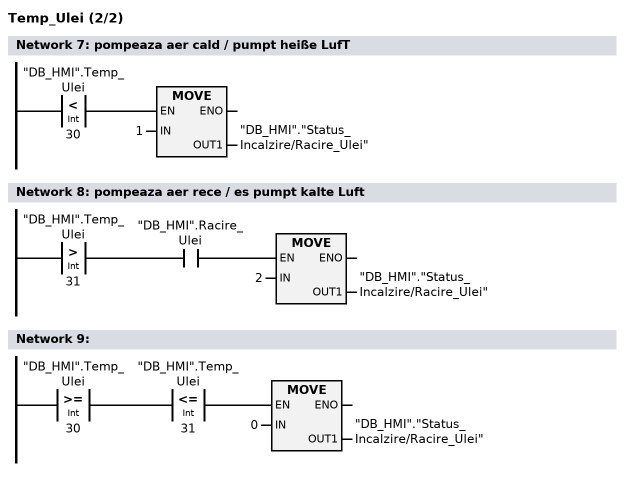
   RUNG wire#powerrail
      { S7_Templates := "SrcType := Int" } LT_Contact(in1 := "DB_HMI".Temp_Ulei, in2 := 30)
      { S7_GenerateENO := "TRUE" } Move(in := 1, out1 => "DB_HMI"."Status_Incalzire/Racire_Ulei")
   END_RUNG
   // the same network as SCL:
   IF "DB_HMI".Temp_Ulei < 30 THEN "DB_HMI"."Status_Incalzire/Racire_Ulei" := 1; END_IF;
END_REGION

REGION Network 8: pompeaza aer rece / es pumpt kalte Luft
   RUNG wire#powerrail
      { S7_Templates := "SrcType := Int" } GT_Contact(in1 := "DB_HMI".Temp_Ulei, in2 := 31)
      Contact( "DB_HMI".Racire_Ulei )
      { S7_GenerateENO := "TRUE" } Move(in := 2, out1 => "DB_HMI"."Status_Incalzire/Racire_Ulei")
   END_RUNG
   // the same network as SCL:
   IF ("DB_HMI".Temp_Ulei > 31) AND "DB_HMI".Racire_Ulei THEN
       "DB_HMI"."Status_Incalzire/Racire_Ulei" := 2;
   END_IF;
END_REGION

REGION Network 9
   RUNG wire#powerrail
      { S7_Templates := "SrcType := Int" } GE_Contact(in1 := "DB_HMI".Temp_Ulei, in2 := 30)
      { S7_Templates := "SrcType := Int" } LE_Contact(in1 := "DB_HMI".Temp_Ulei, in2 := 31)
      { S7_GenerateENO := "TRUE" } Move(in := 0, out1 => "DB_HMI"."Status_Incalzire/Racire_Ulei")
   END_RUNG
   // the same network as SCL:
   IF ("DB_HMI".Temp_Ulei >= 30) AND ("DB_HMI".Temp_Ulei <= 31) THEN
       "DB_HMI"."Status_Incalzire/Racire_Ulei" := 0;
   END_IF;
END_REGION
END_FUNCTION

FUNCTION "Ventilator" : Void   // FC6, LAD
{ S7_Optimized_Access := 'FALSE' }
VERSION : 0.1
BEGIN

REGION Network 1: animatie racire ulei / Ölkühlungsanimation
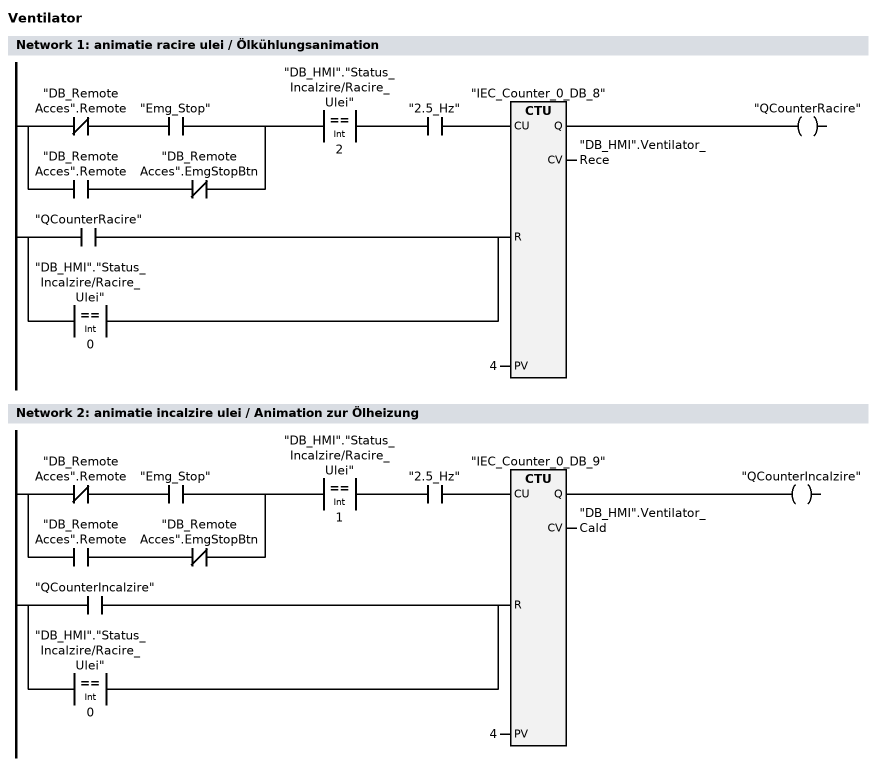
   "IEC_Counter_0_DB_8".CTU(CU := ((NOT "DB_RemoteAcces".Remote AND "Emg_Stop") OR ("DB_RemoteAcces".Remote AND NOT "DB_RemoteAcces".EmgStopBtn)) AND ("DB_HMI"."Status_Incalzire/Racire_Ulei" = 2) AND "2.5_Hz",
                           R := "QCounterRacire" OR ("DB_HMI"."Status_Incalzire/Racire_Ulei" = 0),
                           PV := 4,
                           CV => "DB_HMI".Ventilator_Rece);
   "QCounterRacire" := "IEC_Counter_0_DB_8".Q;
END_REGION

REGION Network 2: animatie incalzire ulei / Animation zur Ölheizung
   "IEC_Counter_0_DB_9".CTU(CU := ((NOT "DB_RemoteAcces".Remote AND "Emg_Stop") OR ("DB_RemoteAcces".Remote AND NOT "DB_RemoteAcces".EmgStopBtn)) AND ("DB_HMI"."Status_Incalzire/Racire_Ulei" = 1) AND "2.5_Hz",
                           R := "QCounterIncalzire" OR ("DB_HMI"."Status_Incalzire/Racire_Ulei" = 0),
                           PV := 4,
                           CV => "DB_HMI".Ventilator_Cald);
   "QCounterIncalzire" := "IEC_Counter_0_DB_9".Q;
END_REGION
END_FUNCTION

FUNCTION "StatusPompe" : Void   // FC19, LAD
{ S7_Optimized_Access := 'FALSE' }
VERSION : 0.1
BEGIN

REGION Network 1
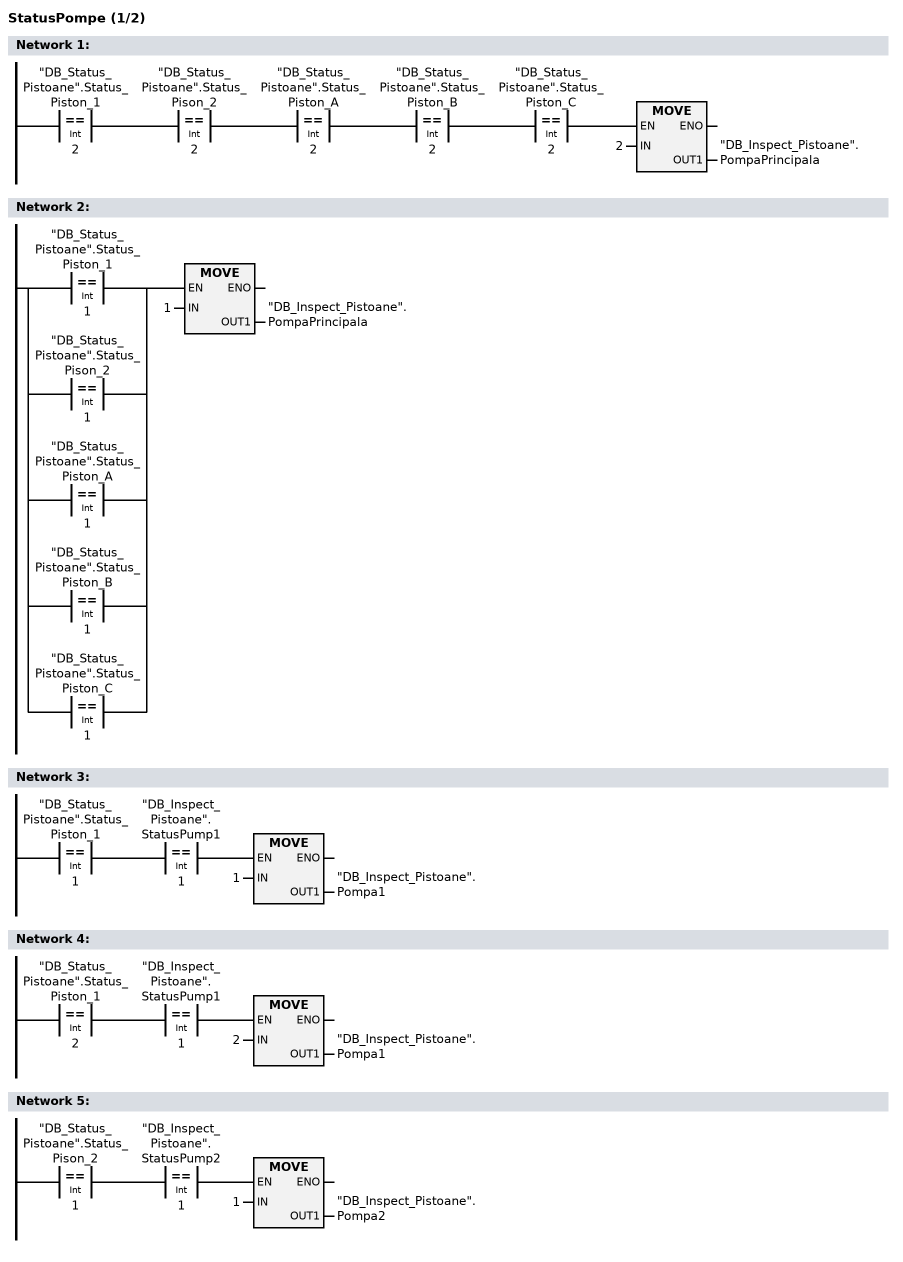
   RUNG wire#powerrail
      { S7_Templates := "SrcType := Int" } EQ_Contact(in1 := "DB_Status_Pistoane".Status_Piston_1, in2 := 2)
      { S7_Templates := "SrcType := Int" } EQ_Contact(in1 := "DB_Status_Pistoane".Status_Pison_2, in2 := 2)
      { S7_Templates := "SrcType := Int" } EQ_Contact(in1 := "DB_Status_Pistoane".Status_Piston_A, in2 := 2)
      { S7_Templates := "SrcType := Int" } EQ_Contact(in1 := "DB_Status_Pistoane".Status_Piston_B, in2 := 2)
      { S7_Templates := "SrcType := Int" } EQ_Contact(in1 := "DB_Status_Pistoane".Status_Piston_C, in2 := 2)
      { S7_GenerateENO := "TRUE" } Move(in := 2, out1 => "DB_Inspect_Pistoane".PompaPrincipala)
   END_RUNG
   // the same network as SCL:
   IF ("DB_Status_Pistoane".Status_Piston_1 = 2) AND ("DB_Status_Pistoane".Status_Pison_2 = 2) AND ("DB_Status_Pistoane".Status_Piston_A = 2) AND ("DB_Status_Pistoane".Status_Piston_B = 2) AND ("DB_Status_Pistoane".Status_Piston_C = 2) THEN
       "DB_Inspect_Pistoane".PompaPrincipala := 2;
   END_IF;
END_REGION

REGION Network 2
   RUNG wire#powerrail
      { S7_Templates := "SrcType := Int" } EQ_Contact(in1 := "DB_Status_Pistoane".Status_Piston_1, in2 := 1)
      wire#w1
      { S7_GenerateENO := "TRUE" } Move(in := 1, out1 => "DB_Inspect_Pistoane".PompaPrincipala)
   END_RUNG
   RUNG wire#powerrail
      { S7_Templates := "SrcType := Int" } EQ_Contact(in1 := "DB_Status_Pistoane".Status_Pison_2, in2 := 1)
   END_RUNG wire#w1
   RUNG wire#powerrail
      { S7_Templates := "SrcType := Int" } EQ_Contact(in1 := "DB_Status_Pistoane".Status_Piston_A, in2 := 1)
   END_RUNG wire#w1
   RUNG wire#powerrail
      { S7_Templates := "SrcType := Int" } EQ_Contact(in1 := "DB_Status_Pistoane".Status_Piston_B, in2 := 1)
   END_RUNG wire#w1
   RUNG wire#powerrail
      { S7_Templates := "SrcType := Int" } EQ_Contact(in1 := "DB_Status_Pistoane".Status_Piston_C, in2 := 1)
   END_RUNG wire#w1
   // the same network as SCL:
   IF ("DB_Status_Pistoane".Status_Piston_1 = 1) OR ("DB_Status_Pistoane".Status_Pison_2 = 1) OR ("DB_Status_Pistoane".Status_Piston_A = 1) OR ("DB_Status_Pistoane".Status_Piston_B = 1) OR ("DB_Status_Pistoane".Status_Piston_C = 1) THEN
       "DB_Inspect_Pistoane".PompaPrincipala := 1;
   END_IF;
END_REGION

REGION Network 3
   RUNG wire#powerrail
      { S7_Templates := "SrcType := Int" } EQ_Contact(in1 := "DB_Status_Pistoane".Status_Piston_1, in2 := 1)
      { S7_Templates := "SrcType := Int" } EQ_Contact(in1 := "DB_Inspect_Pistoane".StatusPump1, in2 := 1)
      { S7_GenerateENO := "TRUE" } Move(in := 1, out1 => "DB_Inspect_Pistoane".Pompa1)
   END_RUNG
   // the same network as SCL:
   IF ("DB_Status_Pistoane".Status_Piston_1 = 1) AND ("DB_Inspect_Pistoane".StatusPump1 = 1) THEN
       "DB_Inspect_Pistoane".Pompa1 := 1;
   END_IF;
END_REGION

REGION Network 4
   RUNG wire#powerrail
      { S7_Templates := "SrcType := Int" } EQ_Contact(in1 := "DB_Status_Pistoane".Status_Piston_1, in2 := 2)
      { S7_Templates := "SrcType := Int" } EQ_Contact(in1 := "DB_Inspect_Pistoane".StatusPump1, in2 := 1)
      { S7_GenerateENO := "TRUE" } Move(in := 2, out1 => "DB_Inspect_Pistoane".Pompa1)
   END_RUNG
   // the same network as SCL:
   IF ("DB_Status_Pistoane".Status_Piston_1 = 2) AND ("DB_Inspect_Pistoane".StatusPump1 = 1) THEN
       "DB_Inspect_Pistoane".Pompa1 := 2;
   END_IF;
END_REGION

REGION Network 5
   RUNG wire#powerrail
      { S7_Templates := "SrcType := Int" } EQ_Contact(in1 := "DB_Status_Pistoane".Status_Pison_2, in2 := 1)
      { S7_Templates := "SrcType := Int" } EQ_Contact(in1 := "DB_Inspect_Pistoane".StatusPump2, in2 := 1)
      { S7_GenerateENO := "TRUE" } Move(in := 1, out1 => "DB_Inspect_Pistoane".Pompa2)
   END_RUNG
   // the same network as SCL:
   IF ("DB_Status_Pistoane".Status_Pison_2 = 1) AND ("DB_Inspect_Pistoane".StatusPump2 = 1) THEN
       "DB_Inspect_Pistoane".Pompa2 := 1;
   END_IF;
END_REGION

REGION Network 6
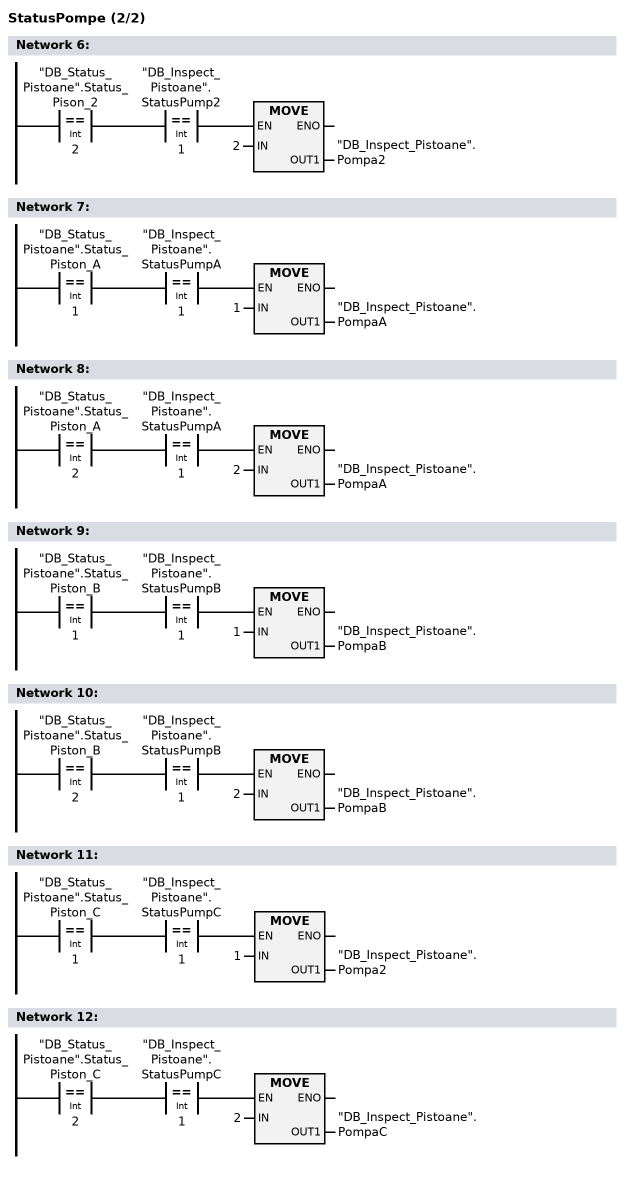
   RUNG wire#powerrail
      { S7_Templates := "SrcType := Int" } EQ_Contact(in1 := "DB_Status_Pistoane".Status_Pison_2, in2 := 2)
      { S7_Templates := "SrcType := Int" } EQ_Contact(in1 := "DB_Inspect_Pistoane".StatusPump2, in2 := 1)
      { S7_GenerateENO := "TRUE" } Move(in := 2, out1 => "DB_Inspect_Pistoane".Pompa2)
   END_RUNG
   // the same network as SCL:
   IF ("DB_Status_Pistoane".Status_Pison_2 = 2) AND ("DB_Inspect_Pistoane".StatusPump2 = 1) THEN
       "DB_Inspect_Pistoane".Pompa2 := 2;
   END_IF;
END_REGION

REGION Network 7
   RUNG wire#powerrail
      { S7_Templates := "SrcType := Int" } EQ_Contact(in1 := "DB_Status_Pistoane".Status_Piston_A, in2 := 1)
      { S7_Templates := "SrcType := Int" } EQ_Contact(in1 := "DB_Inspect_Pistoane".StatusPumpA, in2 := 1)
      { S7_GenerateENO := "TRUE" } Move(in := 1, out1 => "DB_Inspect_Pistoane".PompaA)
   END_RUNG
   // the same network as SCL:
   IF ("DB_Status_Pistoane".Status_Piston_A = 1) AND ("DB_Inspect_Pistoane".StatusPumpA = 1) THEN
       "DB_Inspect_Pistoane".PompaA := 1;
   END_IF;
END_REGION

REGION Network 8
   RUNG wire#powerrail
      { S7_Templates := "SrcType := Int" } EQ_Contact(in1 := "DB_Status_Pistoane".Status_Piston_A, in2 := 2)
      { S7_Templates := "SrcType := Int" } EQ_Contact(in1 := "DB_Inspect_Pistoane".StatusPumpA, in2 := 1)
      { S7_GenerateENO := "TRUE" } Move(in := 2, out1 => "DB_Inspect_Pistoane".PompaA)
   END_RUNG
   // the same network as SCL:
   IF ("DB_Status_Pistoane".Status_Piston_A = 2) AND ("DB_Inspect_Pistoane".StatusPumpA = 1) THEN
       "DB_Inspect_Pistoane".PompaA := 2;
   END_IF;
END_REGION

REGION Network 9
   RUNG wire#powerrail
      { S7_Templates := "SrcType := Int" } EQ_Contact(in1 := "DB_Status_Pistoane".Status_Piston_B, in2 := 1)
      { S7_Templates := "SrcType := Int" } EQ_Contact(in1 := "DB_Inspect_Pistoane".StatusPumpB, in2 := 1)
      { S7_GenerateENO := "TRUE" } Move(in := 1, out1 => "DB_Inspect_Pistoane".PompaB)
   END_RUNG
   // the same network as SCL:
   IF ("DB_Status_Pistoane".Status_Piston_B = 1) AND ("DB_Inspect_Pistoane".StatusPumpB = 1) THEN
       "DB_Inspect_Pistoane".PompaB := 1;
   END_IF;
END_REGION

REGION Network 10
   RUNG wire#powerrail
      { S7_Templates := "SrcType := Int" } EQ_Contact(in1 := "DB_Status_Pistoane".Status_Piston_B, in2 := 2)
      { S7_Templates := "SrcType := Int" } EQ_Contact(in1 := "DB_Inspect_Pistoane".StatusPumpB, in2 := 1)
      { S7_GenerateENO := "TRUE" } Move(in := 2, out1 => "DB_Inspect_Pistoane".PompaB)
   END_RUNG
   // the same network as SCL:
   IF ("DB_Status_Pistoane".Status_Piston_B = 2) AND ("DB_Inspect_Pistoane".StatusPumpB = 1) THEN
       "DB_Inspect_Pistoane".PompaB := 2;
   END_IF;
END_REGION

REGION Network 11
   RUNG wire#powerrail
      { S7_Templates := "SrcType := Int" } EQ_Contact(in1 := "DB_Status_Pistoane".Status_Piston_C, in2 := 1)
      { S7_Templates := "SrcType := Int" } EQ_Contact(in1 := "DB_Inspect_Pistoane".StatusPumpC, in2 := 1)
      { S7_GenerateENO := "TRUE" } Move(in := 1, out1 => "DB_Inspect_Pistoane".Pompa2)
   END_RUNG
   // the same network as SCL:
   IF ("DB_Status_Pistoane".Status_Piston_C = 1) AND ("DB_Inspect_Pistoane".StatusPumpC = 1) THEN
       "DB_Inspect_Pistoane".Pompa2 := 1;
   END_IF;
END_REGION

REGION Network 12
   RUNG wire#powerrail
      { S7_Templates := "SrcType := Int" } EQ_Contact(in1 := "DB_Status_Pistoane".Status_Piston_C, in2 := 2)
      { S7_Templates := "SrcType := Int" } EQ_Contact(in1 := "DB_Inspect_Pistoane".StatusPumpC, in2 := 1)
      { S7_GenerateENO := "TRUE" } Move(in := 2, out1 => "DB_Inspect_Pistoane".PompaC)
   END_RUNG
   // the same network as SCL:
   IF ("DB_Status_Pistoane".Status_Piston_C = 2) AND ("DB_Inspect_Pistoane".StatusPumpC = 1) THEN
       "DB_Inspect_Pistoane".PompaC := 2;
   END_IF;
END_REGION
END_FUNCTION

// folder: Statie Distribuire/Animatii

FUNCTION_BLOCK "Animatie_Banda_1"   // FB2, LAD
{ S7_Optimized_Access := 'FALSE' }
VERSION : 0.1
   VAR_TEMP   // added for the SCL form of the ladder/FBD networks
      _w1 : Bool;
      _w2 : Bool;
   END_VAR
BEGIN

REGION Network 1: ceva
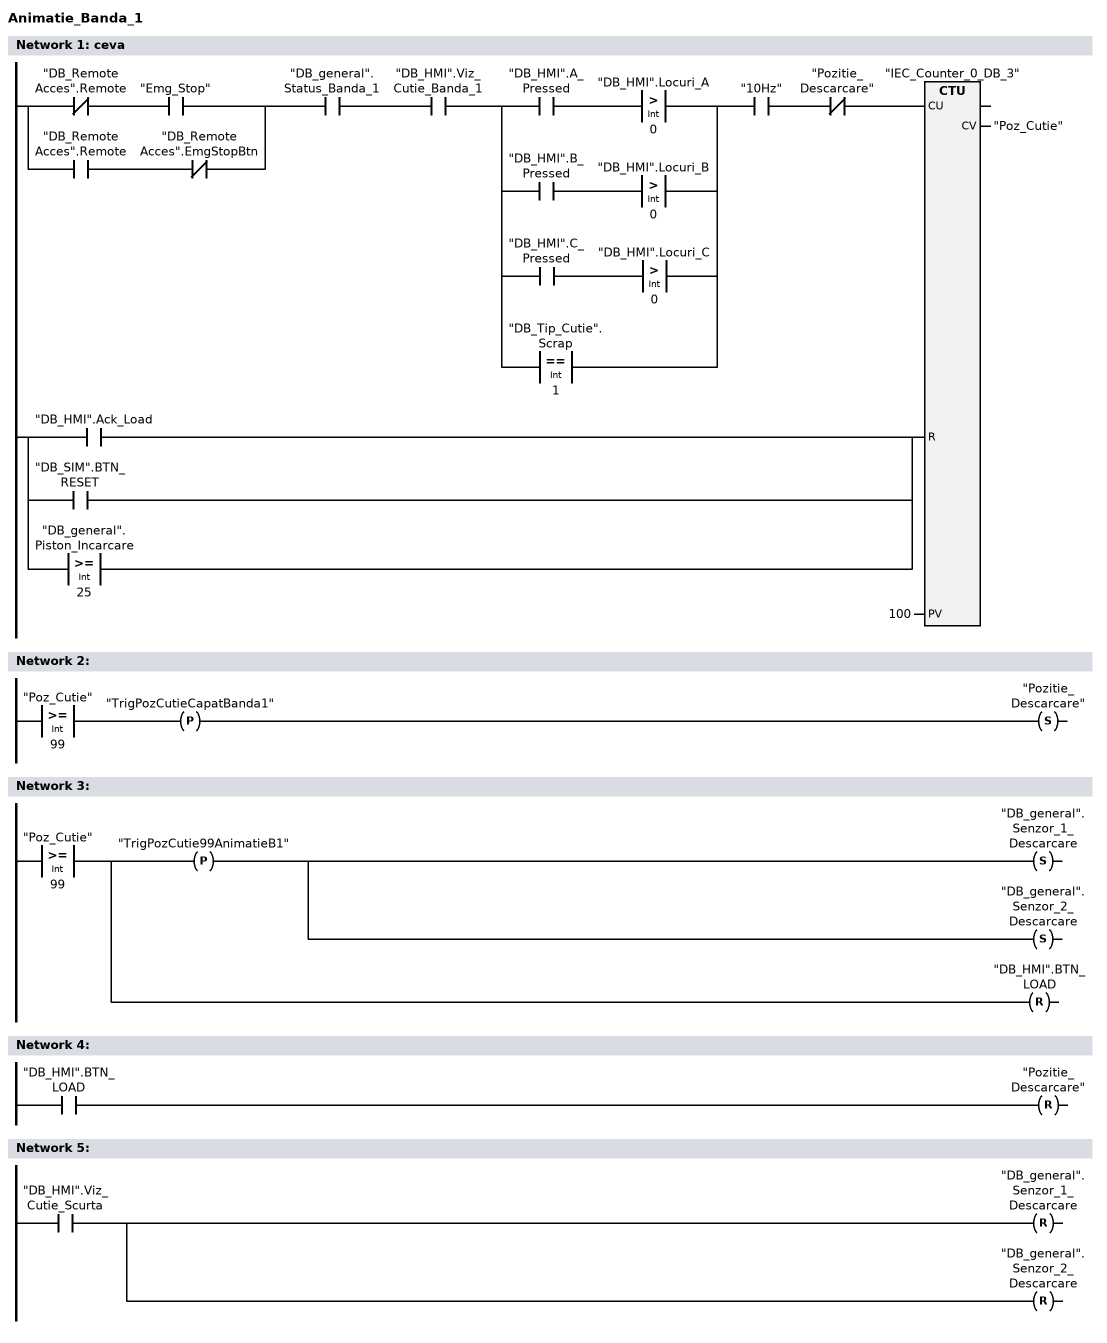
   "IEC_Counter_0_DB_3".CTU(CU := ((NOT "DB_RemoteAcces".Remote AND "Emg_Stop") OR ("DB_RemoteAcces".Remote AND NOT "DB_RemoteAcces".EmgStopBtn)) AND "DB_general".Status_Banda_1 AND "DB_HMI".Viz_Cutie_Banda_1 AND (("DB_HMI".A_Pressed AND ("DB_HMI".Locuri_A > 0)) OR ("DB_HMI".B_Pressed AND ("DB_HMI".Locuri_B > 0)) OR ("DB_HMI".C_Pressed AND ("DB_HMI".Locuri_C > 0)) OR ("DB_Tip_Cutie".Scrap = 1)) AND "10Hz" AND NOT "Pozitie_Descarcare",
                           R := "DB_HMI".Ack_Load OR "DB_SIM".BTN_RESET OR ("DB_general".Piston_Incarcare >= 25),
                           PV := 100,
                           CV => "Poz_Cutie");
END_REGION

REGION Network 2
   RUNG wire#powerrail
      { S7_Templates := "SrcType := Int" } GE_Contact(in1 := "Poz_Cutie", in2 := 99)
      P_Trig( "TrigPozCutieCapatBanda1" )
      S_Coil( "Pozitie_Descarcare" )
   END_RUNG
   // the same network as SCL:
   #_w1 := "Poz_Cutie" >= 99;
   #_w2 := #_w1 AND NOT "TrigPozCutieCapatBanda1";   // rising edge
   "TrigPozCutieCapatBanda1" := #_w1;
   IF #_w2 THEN "Pozitie_Descarcare" := TRUE; END_IF;
END_REGION

REGION Network 3
   RUNG wire#powerrail
      { S7_Templates := "SrcType := Int" } GE_Contact(in1 := "Poz_Cutie", in2 := 99)
      wire#w1
      P_Trig( "TrigPozCutie99AnimatieB1" )
      wire#w2
      S_Coil( "DB_general".Senzor_1_Descarcare )
   END_RUNG
   RUNG wire#w2
      S_Coil( "DB_general".Senzor_2_Descarcare )
   END_RUNG
   RUNG wire#w1
      R_Coil( "DB_HMI".BTN_LOAD )
   END_RUNG
   // the same network as SCL:
   #_w1 := "Poz_Cutie" >= 99;
   #_w2 := #_w1 AND NOT "TrigPozCutie99AnimatieB1";   // rising edge
   "TrigPozCutie99AnimatieB1" := #_w1;
   IF #_w2 THEN
       "DB_general".Senzor_1_Descarcare := TRUE;
       "DB_general".Senzor_2_Descarcare := TRUE;
   END_IF;
   IF #_w1 THEN "DB_HMI".BTN_LOAD := FALSE; END_IF;
END_REGION

REGION Network 4
   RUNG wire#powerrail
      Contact( "DB_HMI".BTN_LOAD )
      R_Coil( "Pozitie_Descarcare" )
   END_RUNG
   // the same network as SCL:
   IF "DB_HMI".BTN_LOAD THEN "Pozitie_Descarcare" := FALSE; END_IF;
END_REGION

REGION Network 5
   RUNG wire#powerrail
      Contact( "DB_HMI".Viz_Cutie_Scurta )
      wire#w1
      R_Coil( "DB_general".Senzor_1_Descarcare )
   END_RUNG
   RUNG wire#w1
      R_Coil( "DB_general".Senzor_2_Descarcare )
   END_RUNG
   // the same network as SCL:
   IF "DB_HMI".Viz_Cutie_Scurta THEN
       "DB_general".Senzor_1_Descarcare := FALSE;
       "DB_general".Senzor_2_Descarcare := FALSE;
   END_IF;
END_REGION
END_FUNCTION_BLOCK

FUNCTION_BLOCK "TranzitieBanda1-Graph"   // FB9, GRAPH
{ S7_Optimized_Access := 'FALSE' }
VERSION : 0.1
   VAR_INPUT
      OFF_SQ : Bool := false;   // Turn sequence off
      INIT_SQ : Bool := false;   // Set sequence to initial state
      ACK_EF : Bool := false;   // Acknowledge all errors and faults
      S_PREV : Bool := false;   // Output previous step in parameter S_NO
      S_NEXT : Bool := false;   // Indicate next step in parameter S_NO
      SW_AUTO : Bool := false;   // Automatic mode
      SW_TAP : Bool := false;   // Semiautomatic/switch with transition
      SW_TOP : Bool := false;   // Semiautomatic/ignore transition
      SW_MAN : Bool := false;   // Manual mode
      S_SEL : Int := 0;   // Select step to be output to S_NO
      S_ON : Bool := false;   // Activate step indicated in S_NO
      S_OFF : Bool := false;   // Deactivate step indicated S_NO
      T_PUSH : Bool := false;   // Enable transition to switch in semi automatic mode
   END_VAR
   VAR_OUTPUT
      S_NO : Int := 0;   // Step number
      S_MORE : Bool := false;   // More steps are available and can be shown in S_NO
      S_ACTIVE : Bool := false;   // Step indicated in S_NO is active
      ERR_FLT : Bool := false;   // Interlock or supervision group error
      AUTO_ON : Bool := false;   // Automatic mode is active
      TAP_ON : Bool := false;   // Semiautomatic mode/step with transition enabled
      TOP_ON : Bool := false;   // Semiautomatic mode/ignore transition enabled
      MAN_ON : Bool := false;   // Manual mode is active
   END_VAR
   VAR
      SWITCH : Array[0..3] of DWord;
      SW_SQTS : Array[0..10] of Byte;
      SW_ADDR : Word := 16#A;
      G7T_0 : GraphTransition;
      G7S_0 : GraphStep;
      PRE_CRIT : Array[0..0] of DWord;
      POST_CRIT : Array[0..0] of DWord;
      TVX : Array[0..12] of Byte;
      TTX : Array[0..12] of Byte;
      TSX : Array[0..2] of Byte;
      S00X : Array[0..2] of Byte;
      SOFFX : Array[0..2] of Byte;
      SONX : Array[0..2] of Byte;
      SAX : Array[0..2] of Byte;
      SERRX : Array[0..11] of Byte;
      SMX : Array[0..11] of Byte;
      S0X : Array[0..11] of Byte;
      S1X : Array[0..11] of Byte;
      S_DISPLAY : Int;   // Internal display of output parameter S_NO
      S_SEL_OLD : Int;   // Previous value in S_SEL
      S_DISPIDX : Byte;   // Index of the step in S_NO
      T_DISPIDX : Byte;   // Index of the transition displayed in T_NO
      MOPEDGE : Struct
         AUTO : Bool := false;
         MAN : Bool := false;
         TAP : Bool := false;
         TOP : Bool := false;
         ACK_S : Bool := false;
         REG_S : Bool := false;
         T_PREV : Bool := false;
         T_NEXT : Bool := false;
         LOCK : Bool := false;
         SUP : Bool := false;
         ACKREQ : Bool := false;
         SSKIP : Bool := false;
         OFF : Bool := false;
         INIT : Bool := false;
         HALT : Bool := false;
         TMS_HALT : Bool := false;
         OPS_ZERO : Bool := false;
         SACT_DISP : Bool := false;
         SEF_DISP : Bool := false;
         SALL_DISP : Bool := false;
         S_PREV : Bool := false;
         S_NEXT : Bool := false;
         S_SELOK : Bool := false;
         S_ON : Bool := false;
         S_OFF : Bool := false;
         T_PUSH : Bool := false;
         REG : Bool := false;
         ACK : Bool := false;
         IL_PERM : Bool := false;
         T_PERM : Bool := false;
         ILP_MAN : Bool := false;
      END_STRUCT;
      MOP : Struct   // Mode
         AUTO : Bool := true;   // Status: automatic mode
         MAN : Bool := false;   // Status: manual mode
         TAP : Bool := false;   // Status: semi automatic/switch with transition
         TOP : Bool := false;   // Status: semi automatic/ignore transition
         ACK_S : Bool := false;   // Request: acknowledge step at parameter S_NO
         REG_S : Bool := false;   // Request: register step indicated in S_NO
         T_PREV : Bool := false;   // Request: output previous valid transition in T_NO
         T_NEXT : Bool := false;   // Request: output next valid transition in T_NO
         LOCK : Bool := true;   // Status: interlocks activated
         SUP : Bool := true;   // Status: supervisions activated
         ACKREQ : Bool := true;   // Status: acknowledgment required
         SSKIP : Bool := false;   // Status: "Skip steps" enabled
         OFF : Bool := false;   // Request: deactivate all steps
         INIT : Bool := true;   // Request: set sequence to initial state
         HALT : Bool := false;   // Status: sequence halted
         TMS_HALT : Bool := false;   // Status: all internal timers held
         OPS_ZERO : Bool := false;   // Status: set all operands processed with N, L, D instructions to 0
         SACT_DISP : Bool := true;   // Status: display active steps only
         SEF_DISP : Bool := false;   // Status: display only steps with errors and disrupted steps
         SALL_DISP : Bool := false;   // Status: display all steps
         S_PREV : Bool := false;   // Request: output previous step to S_NO
         S_NEXT : Bool := false;   // Request: Output next step at S_NO parameter
         S_SELOK : Bool := false;   // Request: output step number from S_SEL to S_NO
         S_ON : Bool := false;   // Request: activate step indicated in S_NO
         S_OFF : Bool := false;   // Request: deactivate step at parameter S_NO
         T_PUSH : Bool := false;   // Request: transition switching enabled
         REG : Bool := false;   // Request: register all interlock and supervision errors
         ACK : Bool := false;   // Request: acknowledge all interlock and supervision errors
         IL_PERM : Bool := false;   // Status: permanent processing of all interlocks
         T_PERM : Bool := false;   // Status: permanent processing of all transitions
         ILP_MAN : Bool := false;   // Status: permanent processing of all interlocks in manual mode
      END_STRUCT;
      TICKS : Struct   // Clock speeds
         DELTA : Time := T#0ms;   // Time difference between cycles
         OLD : Time := T#0ms;   // 10 ms clock counter value in last cycle
         NEW : Time := T#0ms;   // 10 ms clock counter value in this cycle
      END_STRUCT;
      SQ_FLAGS : Struct   // Sequence bit memory
         ERR_FLT : Bool := false;   // Interlock and supervision group error
         ERROR : Bool := false;   // Interlock group error
         FAULT : Bool := false;   // Supervision group error
         RT_FAIL : Bool := false;   // Runtime error
         NO_SNO : Bool := false;   // Requested step number not found
         NF_OFL : Bool := false;   // Overflow: too many ON or OFF requests
         SA_OFL : Bool := false;   // Overflow: too many steps active
         TV_OFL : Bool := false;   // Overflow: too many valid transitions
         MSG_OFL : Bool := false;   // Overflow: not enough system resources for ALARM_S
         NO_SWI : Bool := false;   // Do not switch in this cycle
         CYC_OP : Bool := false;   // Cyclic execution of the sequence after initialization
         AS_MSG : Bool := true;   // Alarms during runtime enabled or disabled by instruction
         AS_SEND : Bool := false;   // Send alarms from WR_USMSG or only enter in diagnostics buffer
         SQ_BUSY : Bool := false;   // Internal edge bit memory for sequence processing
         SA_BUSY : Bool := false;   // Internal edge bit memory for sequence processing
         AS_SIG : Bool := false;   // Edge bit memory for alarms from Alarm_S and Alarm_SQ
      END_STRUCT;
      S_PTR : DWord := 16#940;
      S_PTR2 : DWord := 16#0;
      S_PTR3 : DWord := 16#1720;
      S_PTR4 : DWord := 16#16C0;
      T_PTR : DWord := 16#1660;
      C_AR2 : DWord := 16#0;
      M_FBDB : DWord := 16#90000;
      M_SNO : Word := 16#0;
      M_EVID : Word := 16#0;
      M_EVIL : C_Alarm_s;
      M_EVSV : C_Alarm_s;
      M_EV : DWord := 16#15A0;
      CRIT : Array[0..31] of Bool;
      S_START : Byte := 16#0;
      S_IDX : Byte := 16#0;
      S_INT : Int := 72;
      S_TMP : Byte := 16#0;
      T_START : Byte := 16#0;
      T_IDX : Byte := 16#0;
      T_TMP : Byte := 16#0;
      T_TMP2 : Byte := 16#00;
      TV_POT : Byte := 16#06;
      RETURN1 : Byte := 16#0;
      RETURN2 : Byte := 16#0;
      SINI : Array[0..2] of Byte;
      LSTT : Array[0..15] of Byte;
      ATAJ : Array[0..15] of Byte;
      ATAB : Array[0..15] of Byte;
      PSTT : Array[0..15] of Byte;
      NSTT : Array[0..15] of Byte;
      ASSJ : Array[0..10] of Byte;
      ASSB : Array[0..10] of Byte;
      PTTS : Array[0..10] of Byte;
      NTTS : Array[0..10] of Byte;
      PRE_CNT : Word := 16#1;
      POST_CNT : Word := 16#1;
      ADR_COND : Word := 16#0;
      MAX_TVAL : Byte := 16#B;
      MAX_SACT : Byte := 16#1;
      MAX_CRIT : Byte := 16#4;
      T_CNT : Byte := 16#F;
      SUP_CNT : Byte := 16#0;
      LOCK_CNT : Byte := 16#0;
      S_CNT : Byte := 16#A;
      SQ_CNT : Byte := 16#1;
      PRS_INPAR : DWord := 16#E000FEC8;
      PRS_OUTPAR : DWord := 16#E000800F;
      GC_FLAGS : Struct
         T_MACH : Byte := 16#EB;
         COND_ED : Byte := 16#E3;
         W_LEVEL : Byte := 16#D5;
         FB_IF : Byte := 16#FA;
         AS_MSG : Word := 16#404;
         SSB : Word := 16#108;
         DILG : Word := 16#3F4;
         ADDR_T0 : Word := 16#28;
         CRIT_AVAIL : Bool := false;
         SSKIP_AVAIL : Bool := true;
         SSKIP_ON : Bool := false;
         ACK_REQ : Bool := true;
         SYNC_AVAIL : Bool := true;
         ILP_MAN : Bool := false;
         SWM_LOCKED : Bool := false;
         SAVE_SW : Bool := true;
      END_STRUCT;
      G7_FBMARK : Byte := 16#3C;
      G7_RELEASE : Byte := 16#3C;
      G7_ID2 : Byte := 16#37;
      G7_ID1 : Byte := 16#47;
   END_VAR
   // SW_SQTS[0] := 16#A;
   // TVX[0] := 16#1;
   // TTX[0] := 16#1;
   // TSX[0] := 16#1;
   // S00X[0] := 16#1;
   // SOFFX[0] := 16#1;
   // SONX[0] := 16#1;
   // SAX[0] := 16#1;
   // SERRX[0] := 16#1;
   // SMX[0] := 16#1;
   // S0X[0] := 16#1;
   // S1X[0] := 16#1;
   // SINI[0] := 16#2;
   // SINI[1] := 16#1;
   // SINI[2] := 0;
   // LSTT[0] := 0;
   // LSTT[1] := 0;
   // LSTT[2] := 0;
   // LSTT[3] := 0;
   // ATAJ[0] := 0;
   // ATAJ[1] := 16#1;
   // ATAJ[2] := 16#2;
   // ATAJ[3] := 16#3;
   // ATAB[0] := 0;
   // ATAB[1] := 16#6;
   // ATAB[2] := 16#9;
   // ATAB[3] := 16#8;
   // PSTT[0] := 0;
   // PSTT[1] := 16#1;
   // PSTT[2] := 16#2;
   // PSTT[3] := 16#3;
   // NSTT[0] := 16#1;
   // NSTT[1] := 16#2;
   // NSTT[2] := 16#3;
   // ASSJ[0] := 0;
   // ASSJ[1] := 16#1;
   // ASSJ[2] := 16#2;
   // ASSJ[3] := 16#3;
   // ASSB[0] := 0;
   // ASSB[1] := 16#1;
   // ASSB[2] := 16#2;
   // ASSB[3] := 16#3;
   // PTTS[0] := 0;
   // PTTS[2] := 16#1;
   // PTTS[3] := 16#2;
   // NTTS[0] := 0;
   // NTTS[1] := 16#1;
   // NTTS[2] := 16#2;
   // NTTS[3] := 16#3;
   // NSTT[3] := 16#4;
   // PSTT[5] := 16#5;
   // ATAB[5] := 16#D;
   // NSTT[5] := 16#1;
   // NSTT[4] := 16#5;
   // NTTS[5] := 16#5;
   // PTTS[5] := 16#4;
   // ASSB[5] := 16#5;
   // ASSJ[5] := 16#5;
   // ATAJ[5] := 16#5;
   // LSTT[5] := 16#1;
   // NTTS[4] := 16#4;
   // PTTS[4] := 16#3;
   // ASSB[4] := 16#4;
   // ASSJ[4] := 16#4;
   // PSTT[4] := 16#4;
   // ATAB[4] := 16#B;
   // ATAJ[4] := 16#4;
   // LSTT[4] := 0;
   // SW_SQTS[2] := 16#1;
   // SW_SQTS[3] := 16#2;
   // SW_SQTS[4] := 16#3;
   // SW_SQTS[5] := 16#4;
   // SW_SQTS[6] := 16#5;
   // SW_SQTS[7] := 16#6;
   // LSTT[6] := 0;
   // LSTT[7] := 16#1;
   // LSTT[8] := 0;
   // LSTT[9] := 0;
   // ATAJ[6] := 16#6;
   // ATAJ[7] := 16#7;
   // ATAJ[8] := 16#8;
   // ATAJ[9] := 16#9;
   // ATAB[6] := 16#1;
   // ATAB[7] := 16#7;
   // ATAB[8] := 16#3;
   // ATAB[9] := 16#2;
   // PSTT[6] := 16#1;
   // PSTT[7] := 16#6;
   // PSTT[8] := 16#3;
   // PSTT[9] := 16#2;
   // NSTT[6] := 16#6;
   // NSTT[7] := 16#1;
   // NSTT[8] := 16#8;
   // NSTT[9] := 16#7;
   // ASSJ[6] := 16#6;
   // ASSJ[7] := 16#7;
   // ASSB[6] := 16#6;
   // ASSB[7] := 16#7;
   // PTTS[6] := 16#6;
   // PTTS[7] := 16#9;
   // NTTS[6] := 16#7;
   // NTTS[7] := 16#A;
   // SW_SQTS[8] := 16#7;
   // SW_SQTS[9] := 16#8;
   // SW_SQTS[10] := 16#9;
   // LSTT[10] := 16#1;
   // LSTT[11] := 0;
   // LSTT[12] := 16#1;
   // LSTT[13] := 0;
   // LSTT[14] := 16#1;
   // LSTT[15] := 16#1;
   // ATAJ[10] := 16#A;
   // ATAJ[11] := 16#B;
   // ATAJ[12] := 16#C;
   // ATAJ[13] := 16#D;
   // ATAJ[14] := 16#E;
   // ATAJ[15] := 16#F;
   // ATAB[10] := 16#A;
   // ATAB[11] := 16#4;
   // ATAB[12] := 16#C;
   // ATAB[13] := 16#5;
   // ATAB[14] := 16#E;
   // ATAB[15] := 16#F;
   // PSTT[10] := 16#7;
   // PSTT[11] := 16#4;
   // PSTT[12] := 16#8;
   // PSTT[13] := 16#5;
   // PSTT[14] := 16#9;
   // PSTT[15] := 16#A;
   // NSTT[10] := 16#1;
   // NSTT[11] := 16#9;
   // NSTT[12] := 16#1;
   // NSTT[13] := 16#A;
   // NSTT[14] := 16#1;
   // NSTT[15] := 16#1;
   // ASSJ[8] := 16#8;
   // ASSJ[9] := 16#9;
   // ASSJ[10] := 16#A;
   // ASSB[8] := 16#8;
   // ASSB[9] := 16#9;
   // ASSB[10] := 16#A;
   // PTTS[8] := 16#8;
   // PTTS[9] := 16#B;
   // PTTS[10] := 16#D;
   // NTTS[8] := 16#C;
   // NTTS[9] := 16#E;
   // NTTS[10] := 16#F;
BEGIN
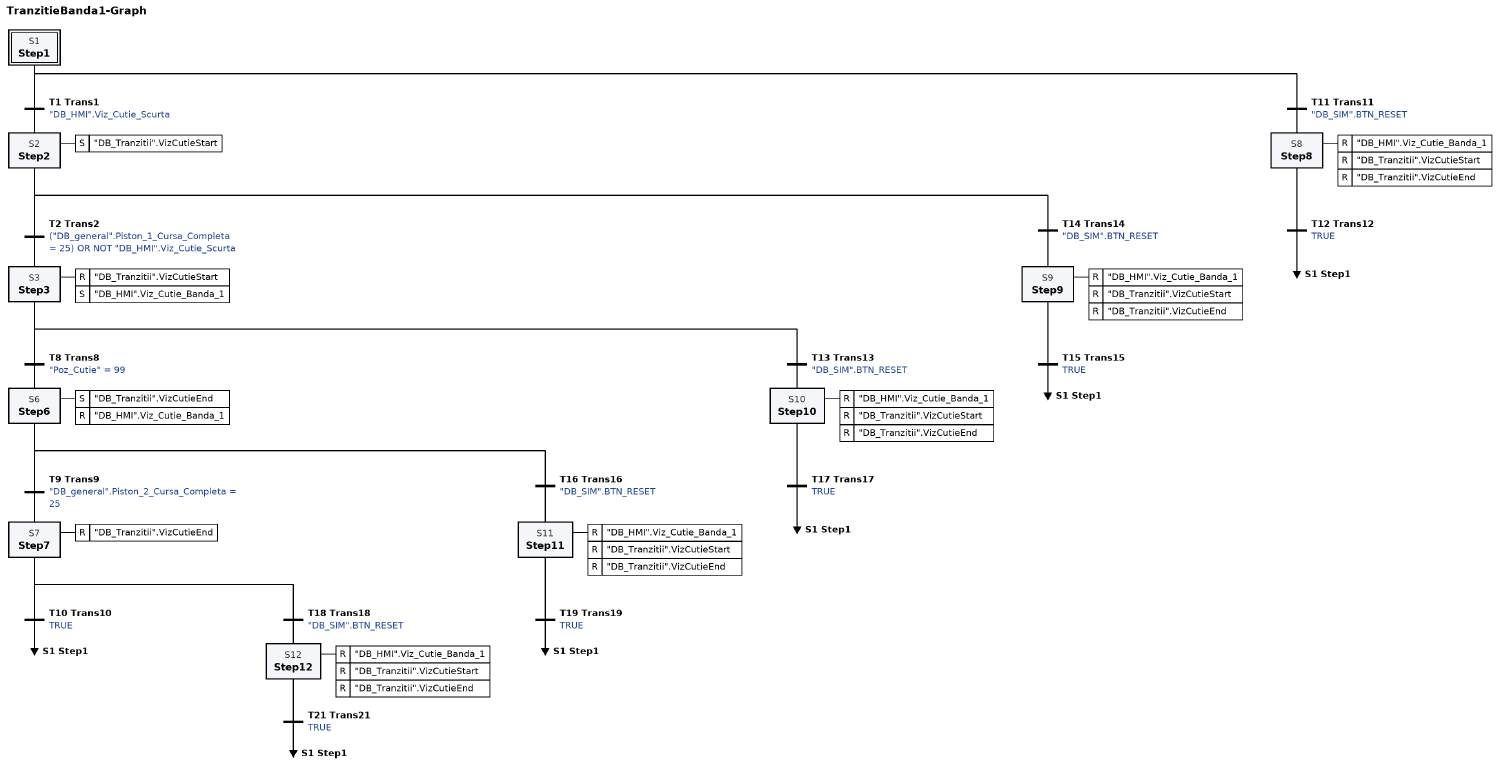
   // sequencer 1
   INITIAL_STEP Step1:   // S1
   END_STEP
   TRANSITION Trans1 FROM Step1 TO Step2   // T1
      := "DB_HMI".Viz_Cutie_Scurta;
   END_TRANSITION
   TRANSITION Trans11 FROM Step1 TO Step8   // T11
      := "DB_SIM".BTN_RESET;
   END_TRANSITION
   STEP Step2:   // S2
              S    "DB_Tranzitii".VizCutieStart
   END_STEP
   TRANSITION Trans2 FROM Step2 TO Step3   // T2
      := ("DB_general".Piston_1_Cursa_Completa = 25) OR NOT "DB_HMI".Viz_Cutie_Scurta;
   END_TRANSITION
   TRANSITION Trans14 FROM Step2 TO Step9   // T14
      := "DB_SIM".BTN_RESET;
   END_TRANSITION
   STEP Step3:   // S3
              R    "DB_Tranzitii".VizCutieStart
              S    "DB_HMI".Viz_Cutie_Banda_1
   END_STEP
   TRANSITION Trans8 FROM Step3 TO Step6   // T8
      := "Poz_Cutie" = 99;
   END_TRANSITION
   TRANSITION Trans13 FROM Step3 TO Step10   // T13
      := "DB_SIM".BTN_RESET;
   END_TRANSITION
   STEP Step6:   // S6
              S    "DB_Tranzitii".VizCutieEnd
              R    "DB_HMI".Viz_Cutie_Banda_1
   END_STEP
   TRANSITION Trans9 FROM Step6 TO Step7   // T9
      := "DB_general".Piston_2_Cursa_Completa = 25;
   END_TRANSITION
   TRANSITION Trans16 FROM Step6 TO Step11   // T16
      := "DB_SIM".BTN_RESET;
   END_TRANSITION
   STEP Step7:   // S7
              R    "DB_Tranzitii".VizCutieEnd
   END_STEP
   TRANSITION Trans10 FROM Step7 TO Step1   // T10, jump
      := TRUE;
   END_TRANSITION
   TRANSITION Trans18 FROM Step7 TO Step12   // T18
      := "DB_SIM".BTN_RESET;
   END_TRANSITION
   STEP Step8:   // S8
              R    "DB_HMI".Viz_Cutie_Banda_1
              R    "DB_Tranzitii".VizCutieStart
              R    "DB_Tranzitii".VizCutieEnd
   END_STEP
   TRANSITION Trans12 FROM Step8 TO Step1   // T12, jump
      := TRUE;
   END_TRANSITION
   STEP Step10:   // S10
              R    "DB_HMI".Viz_Cutie_Banda_1
              R    "DB_Tranzitii".VizCutieStart
              R    "DB_Tranzitii".VizCutieEnd
   END_STEP
   TRANSITION Trans17 FROM Step10 TO Step1   // T17, jump
      := TRUE;
   END_TRANSITION
   STEP Step9:   // S9
              R    "DB_HMI".Viz_Cutie_Banda_1
              R    "DB_Tranzitii".VizCutieStart
              R    "DB_Tranzitii".VizCutieEnd
   END_STEP
   TRANSITION Trans15 FROM Step9 TO Step1   // T15, jump
      := TRUE;
   END_TRANSITION
   STEP Step11:   // S11
              R    "DB_HMI".Viz_Cutie_Banda_1
              R    "DB_Tranzitii".VizCutieStart
              R    "DB_Tranzitii".VizCutieEnd
   END_STEP
   TRANSITION Trans19 FROM Step11 TO Step1   // T19, jump
      := TRUE;
   END_TRANSITION
   STEP Step12:   // S12
              R    "DB_HMI".Viz_Cutie_Banda_1
              R    "DB_Tranzitii".VizCutieStart
              R    "DB_Tranzitii".VizCutieEnd
   END_STEP
   TRANSITION Trans21 FROM Step12 TO Step1   // T21, jump
      := TRUE;
   END_TRANSITION
END_FUNCTION_BLOCK

FUNCTION_BLOCK "Animatie_Piston_1"   // FB10, LAD
{ S7_Optimized_Access := 'FALSE' }
VERSION : 0.1
BEGIN

REGION Network 1
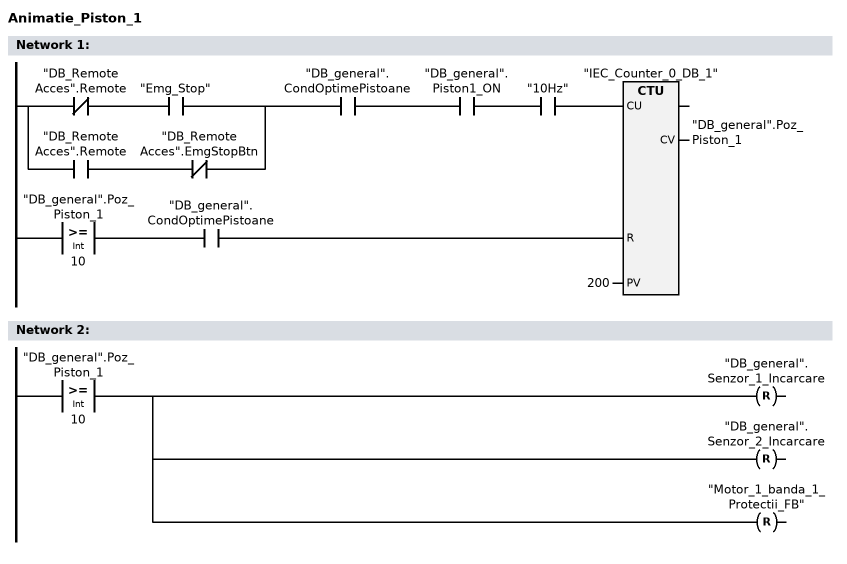
   "IEC_Counter_0_DB_1".CTU(CU := ((NOT "DB_RemoteAcces".Remote AND "Emg_Stop") OR ("DB_RemoteAcces".Remote AND NOT "DB_RemoteAcces".EmgStopBtn)) AND "DB_general".CondOptimePistoane AND "DB_general".Piston1_ON AND "10Hz",
                           R := ("DB_general".Poz_Piston_1 >= 10) AND "DB_general".CondOptimePistoane,
                           PV := 200,
                           CV => "DB_general".Poz_Piston_1);
END_REGION

REGION Network 2
   RUNG wire#powerrail
      { S7_Templates := "SrcType := Int" } GE_Contact(in1 := "DB_general".Poz_Piston_1, in2 := 10)
      wire#w1
      R_Coil( "DB_general".Senzor_1_Incarcare )
   END_RUNG
   RUNG wire#w1
      R_Coil( "DB_general".Senzor_2_Incarcare )
   END_RUNG
   RUNG wire#w1
      R_Coil( "Motor_1_banda_1_Protectii_FB" )
   END_RUNG
   // the same network as SCL:
   IF "DB_general".Poz_Piston_1 >= 10 THEN
       "DB_general".Senzor_1_Incarcare := FALSE;
       "DB_general".Senzor_2_Incarcare := FALSE;
       "Motor_1_banda_1_Protectii_FB" := FALSE;
   END_IF;
END_REGION
END_FUNCTION_BLOCK

FUNCTION_BLOCK "Piston_1_Cursa_Completa"   // FB13, LAD
{ S7_Optimized_Access := 'FALSE' }